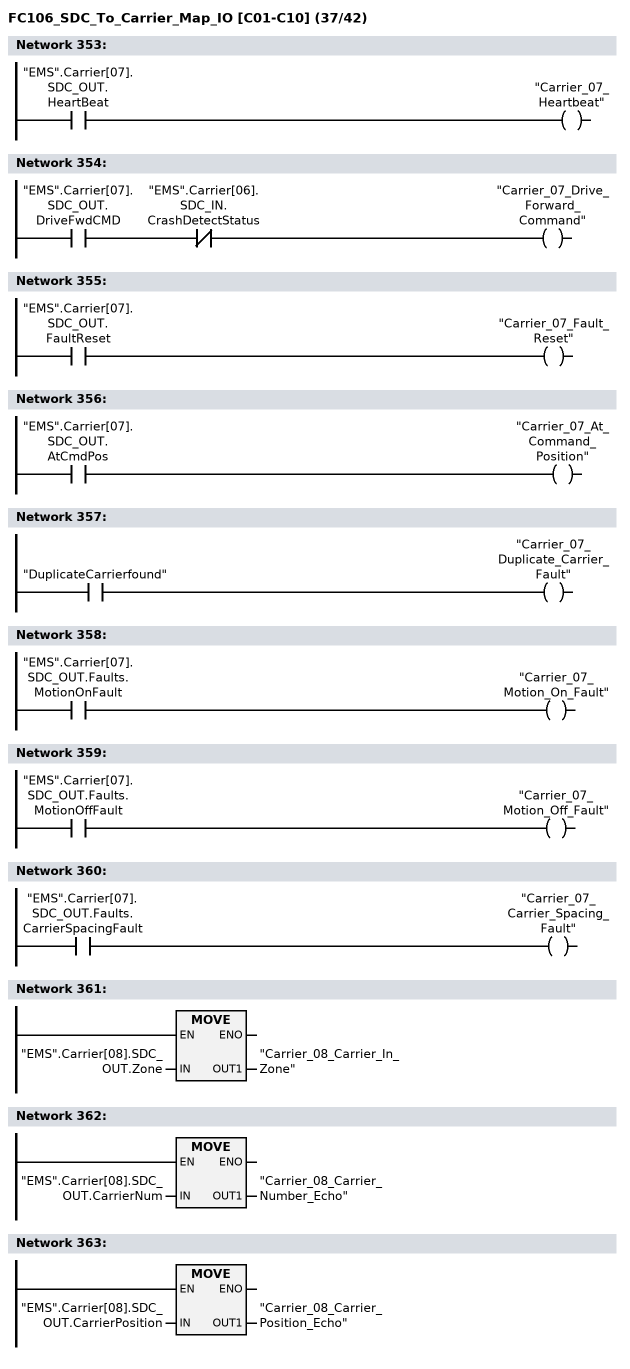
   RUNG wire#powerrail
      Contact( "EMS".Carrier[07].SDC_OUT.HeartBeat )
      Coil( "Carrier_07_Heartbeat" )
   END_RUNG
   // the same network as SCL:
   "Carrier_07_Heartbeat" := "EMS".Carrier[07].SDC_OUT.HeartBeat;
END_REGION

REGION Network 354
   RUNG wire#powerrail
      Contact( "EMS".Carrier[07].SDC_OUT.DriveFwdCMD )
      I_Contact( "EMS".Carrier[06].SDC_IN.CrashDetectStatus )
      Coil( "Carrier_07_Drive_Forward_Command" )
   END_RUNG
   // the same network as SCL:
   "Carrier_07_Drive_Forward_Command" := "EMS".Carrier[07].SDC_OUT.DriveFwdCMD AND NOT "EMS".Carrier[06].SDC_IN.CrashDetectStatus;
END_REGION

REGION Network 355
   RUNG wire#powerrail
      Contact( "EMS".Carrier[07].SDC_OUT.FaultReset )
      Coil( "Carrier_07_Fault_Reset" )
   END_RUNG
   // the same network as SCL:
   "Carrier_07_Fault_Reset" := "EMS".Carrier[07].SDC_OUT.FaultReset;
END_REGION

REGION Network 356
   RUNG wire#powerrail
      Contact( "EMS".Carrier[07].SDC_OUT.AtCmdPos )
      Coil( "Carrier_07_At_Command_Position" )
   END_RUNG
   // the same network as SCL:
   "Carrier_07_At_Command_Position" := "EMS".Carrier[07].SDC_OUT.AtCmdPos;
END_REGION

REGION Network 357
   RUNG wire#powerrail
      Contact( "DuplicateCarrierfound" )
      Coil( "Carrier_07_Duplicate_Carrier_Fault" )
   END_RUNG
   // the same network as SCL:
   "Carrier_07_Duplicate_Carrier_Fault" := "DuplicateCarrierfound";
END_REGION

REGION Network 358
   RUNG wire#powerrail
      Contact( "EMS".Carrier[07].SDC_OUT.Faults.MotionOnFault )
      Coil( "Carrier_07_Motion_On_Fault" )
   END_RUNG
   // the same network as SCL:
   "Carrier_07_Motion_On_Fault" := "EMS".Carrier[07].SDC_OUT.Faults.MotionOnFault;
END_REGION

REGION Network 359
   RUNG wire#powerrail
      Contact( "EMS".Carrier[07].SDC_OUT.Faults.MotionOffFault )
      Coil( "Carrier_07_Motion_Off_Fault" )
   END_RUNG
   // the same network as SCL:
   "Carrier_07_Motion_Off_Fault" := "EMS".Carrier[07].SDC_OUT.Faults.MotionOffFault;
END_REGION

REGION Network 360
   RUNG wire#powerrail
      Contact( "EMS".Carrier[07].SDC_OUT.Faults.CarrierSpacingFault )
      Coil( "Carrier_07_Carrier_Spacing_Fault" )
   END_RUNG
   // the same network as SCL:
   "Carrier_07_Carrier_Spacing_Fault" := "EMS".Carrier[07].SDC_OUT.Faults.CarrierSpacingFault;
END_REGION

REGION Network 361
   RUNG wire#powerrail
      Move(in := "EMS".Carrier[08].SDC_OUT.Zone, out1 => "Carrier_08_Carrier_In_Zone")
   END_RUNG
   // the same network as SCL:
   "Carrier_08_Carrier_In_Zone" := "EMS".Carrier[08].SDC_OUT.Zone;
END_REGION

REGION Network 362
   RUNG wire#powerrail
      Move(in := "EMS".Carrier[08].SDC_OUT.CarrierNum, out1 => "Carrier_08_Carrier_Number_Echo")
   END_RUNG
   // the same network as SCL:
   "Carrier_08_Carrier_Number_Echo" := "EMS".Carrier[08].SDC_OUT.CarrierNum;
END_REGION

REGION Network 363
   RUNG wire#powerrail
      Move(in := "EMS".Carrier[08].SDC_OUT.CarrierPosition, out1 => "Carrier_08_Carrier_Position_Echo")
   END_RUNG
   // the same network as SCL:
   "Carrier_08_Carrier_Position_Echo" := "EMS".Carrier[08].SDC_OUT.CarrierPosition;
END_REGION

REGION Network 364
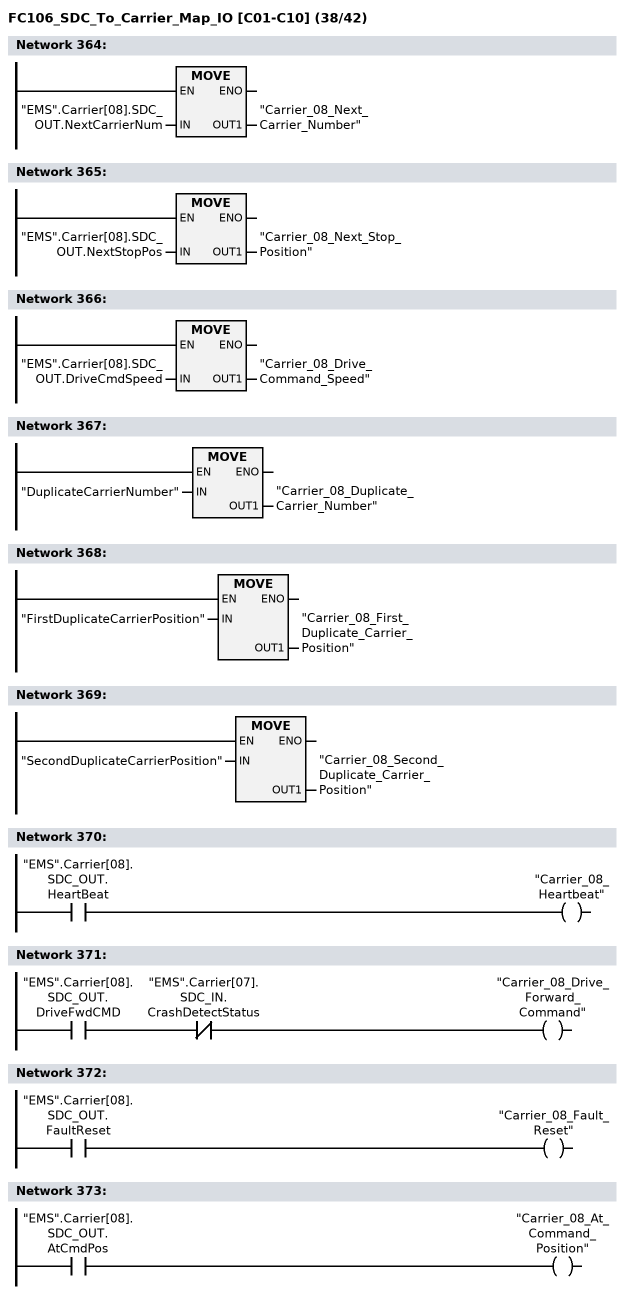
   RUNG wire#powerrail
      Move(in := "EMS".Carrier[08].SDC_OUT.NextCarrierNum, out1 => "Carrier_08_Next_Carrier_Number")
   END_RUNG
   // the same network as SCL:
   "Carrier_08_Next_Carrier_Number" := "EMS".Carrier[08].SDC_OUT.NextCarrierNum;
END_REGION

REGION Network 365
   RUNG wire#powerrail
      Move(in := "EMS".Carrier[08].SDC_OUT.NextStopPos, out1 => "Carrier_08_Next_Stop_Position")
   END_RUNG
   // the same network as SCL:
   "Carrier_08_Next_Stop_Position" := "EMS".Carrier[08].SDC_OUT.NextStopPos;
END_REGION

REGION Network 366
   RUNG wire#powerrail
      Move(in := "EMS".Carrier[08].SDC_OUT.DriveCmdSpeed, out1 => "Carrier_08_Drive_Command_Speed")
   END_RUNG
   // the same network as SCL:
   "Carrier_08_Drive_Command_Speed" := "EMS".Carrier[08].SDC_OUT.DriveCmdSpeed;
END_REGION

REGION Network 367
   RUNG wire#powerrail
      Move(in := "DuplicateCarrierNumber", out1 => "Carrier_08_Duplicate_Carrier_Number")
   END_RUNG
   // the same network as SCL:
   "Carrier_08_Duplicate_Carrier_Number" := "DuplicateCarrierNumber";
END_REGION

REGION Network 368
   RUNG wire#powerrail
      Move(in := "FirstDuplicateCarrierPosition", out1 => "Carrier_08_First_Duplicate_Carrier_Position")
   END_RUNG
   // the same network as SCL:
   "Carrier_08_First_Duplicate_Carrier_Position" := "FirstDuplicateCarrierPosition";
END_REGION

REGION Network 369
   RUNG wire#powerrail
      Move(in := "SecondDuplicateCarrierPosition", out1 => "Carrier_08_Second_Duplicate_Carrier_Position")
   END_RUNG
   // the same network as SCL:
   "Carrier_08_Second_Duplicate_Carrier_Position" := "SecondDuplicateCarrierPosition";
END_REGION

REGION Network 370
   RUNG wire#powerrail
      Contact( "EMS".Carrier[08].SDC_OUT.HeartBeat )
      Coil( "Carrier_08_Heartbeat" )
   END_RUNG
   // the same network as SCL:
   "Carrier_08_Heartbeat" := "EMS".Carrier[08].SDC_OUT.HeartBeat;
END_REGION

REGION Network 371
   RUNG wire#powerrail
      Contact( "EMS".Carrier[08].SDC_OUT.DriveFwdCMD )
      I_Contact( "EMS".Carrier[07].SDC_IN.CrashDetectStatus )
      Coil( "Carrier_08_Drive_Forward_Command" )
   END_RUNG
   // the same network as SCL:
   "Carrier_08_Drive_Forward_Command" := "EMS".Carrier[08].SDC_OUT.DriveFwdCMD AND NOT "EMS".Carrier[07].SDC_IN.CrashDetectStatus;
END_REGION

REGION Network 372
   RUNG wire#powerrail
      Contact( "EMS".Carrier[08].SDC_OUT.FaultReset )
      Coil( "Carrier_08_Fault_Reset" )
   END_RUNG
   // the same network as SCL:
   "Carrier_08_Fault_Reset" := "EMS".Carrier[08].SDC_OUT.FaultReset;
END_REGION

REGION Network 373
   RUNG wire#powerrail
      Contact( "EMS".Carrier[08].SDC_OUT.AtCmdPos )
      Coil( "Carrier_08_At_Command_Position" )
   END_RUNG
   // the same network as SCL:
   "Carrier_08_At_Command_Position" := "EMS".Carrier[08].SDC_OUT.AtCmdPos;
END_REGION

REGION Network 374
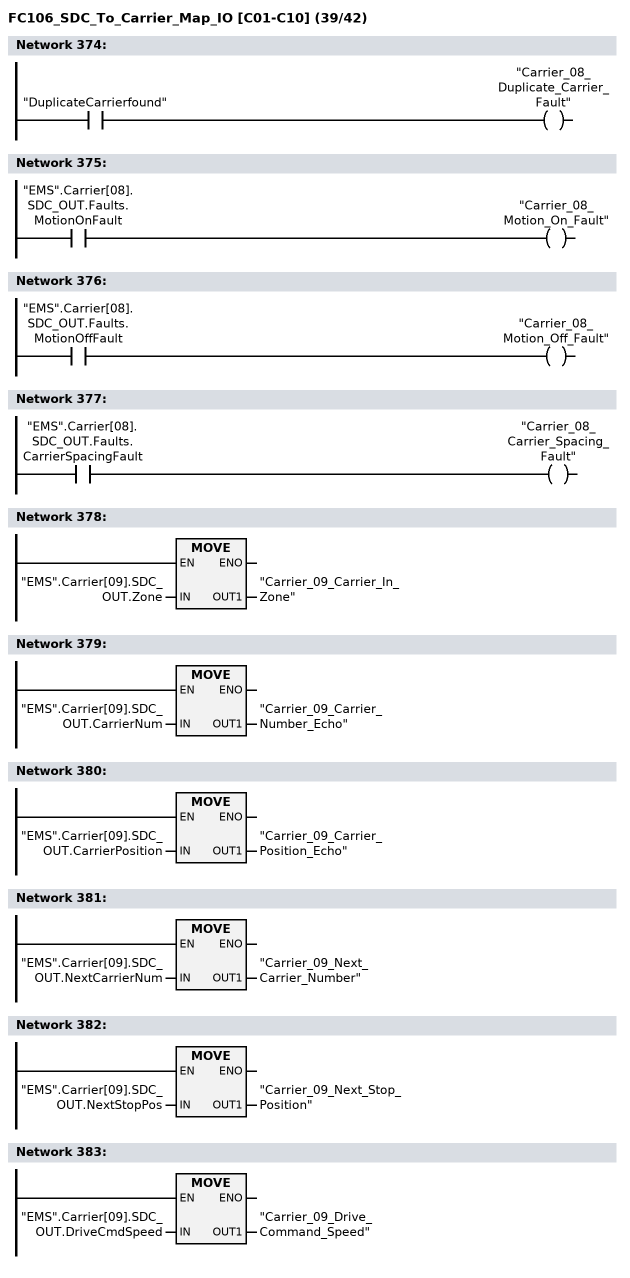
   RUNG wire#powerrail
      Contact( "DuplicateCarrierfound" )
      Coil( "Carrier_08_Duplicate_Carrier_Fault" )
   END_RUNG
   // the same network as SCL:
   "Carrier_08_Duplicate_Carrier_Fault" := "DuplicateCarrierfound";
END_REGION

REGION Network 375
   RUNG wire#powerrail
      Contact( "EMS".Carrier[08].SDC_OUT.Faults.MotionOnFault )
      Coil( "Carrier_08_Motion_On_Fault" )
   END_RUNG
   // the same network as SCL:
   "Carrier_08_Motion_On_Fault" := "EMS".Carrier[08].SDC_OUT.Faults.MotionOnFault;
END_REGION

REGION Network 376
   RUNG wire#powerrail
      Contact( "EMS".Carrier[08].SDC_OUT.Faults.MotionOffFault )
      Coil( "Carrier_08_Motion_Off_Fault" )
   END_RUNG
   // the same network as SCL:
   "Carrier_08_Motion_Off_Fault" := "EMS".Carrier[08].SDC_OUT.Faults.MotionOffFault;
END_REGION

REGION Network 377
   RUNG wire#powerrail
      Contact( "EMS".Carrier[08].SDC_OUT.Faults.CarrierSpacingFault )
      Coil( "Carrier_08_Carrier_Spacing_Fault" )
   END_RUNG
   // the same network as SCL:
   "Carrier_08_Carrier_Spacing_Fault" := "EMS".Carrier[08].SDC_OUT.Faults.CarrierSpacingFault;
END_REGION

REGION Network 378
   RUNG wire#powerrail
      Move(in := "EMS".Carrier[09].SDC_OUT.Zone, out1 => "Carrier_09_Carrier_In_Zone")
   END_RUNG
   // the same network as SCL:
   "Carrier_09_Carrier_In_Zone" := "EMS".Carrier[09].SDC_OUT.Zone;
END_REGION

REGION Network 379
   RUNG wire#powerrail
      Move(in := "EMS".Carrier[09].SDC_OUT.CarrierNum, out1 => "Carrier_09_Carrier_Number_Echo")
   END_RUNG
   // the same network as SCL:
   "Carrier_09_Carrier_Number_Echo" := "EMS".Carrier[09].SDC_OUT.CarrierNum;
END_REGION

REGION Network 380
   RUNG wire#powerrail
      Move(in := "EMS".Carrier[09].SDC_OUT.CarrierPosition, out1 => "Carrier_09_Carrier_Position_Echo")
   END_RUNG
   // the same network as SCL:
   "Carrier_09_Carrier_Position_Echo" := "EMS".Carrier[09].SDC_OUT.CarrierPosition;
END_REGION

REGION Network 381
   RUNG wire#powerrail
      Move(in := "EMS".Carrier[09].SDC_OUT.NextCarrierNum, out1 => "Carrier_09_Next_Carrier_Number")
   END_RUNG
   // the same network as SCL:
   "Carrier_09_Next_Carrier_Number" := "EMS".Carrier[09].SDC_OUT.NextCarrierNum;
END_REGION

REGION Network 382
   RUNG wire#powerrail
      Move(in := "EMS".Carrier[09].SDC_OUT.NextStopPos, out1 => "Carrier_09_Next_Stop_Position")
   END_RUNG
   // the same network as SCL:
   "Carrier_09_Next_Stop_Position" := "EMS".Carrier[09].SDC_OUT.NextStopPos;
END_REGION

REGION Network 383
   RUNG wire#powerrail
      Move(in := "EMS".Carrier[09].SDC_OUT.DriveCmdSpeed, out1 => "Carrier_09_Drive_Command_Speed")
   END_RUNG
   // the same network as SCL:
   "Carrier_09_Drive_Command_Speed" := "EMS".Carrier[09].SDC_OUT.DriveCmdSpeed;
END_REGION

REGION Network 384
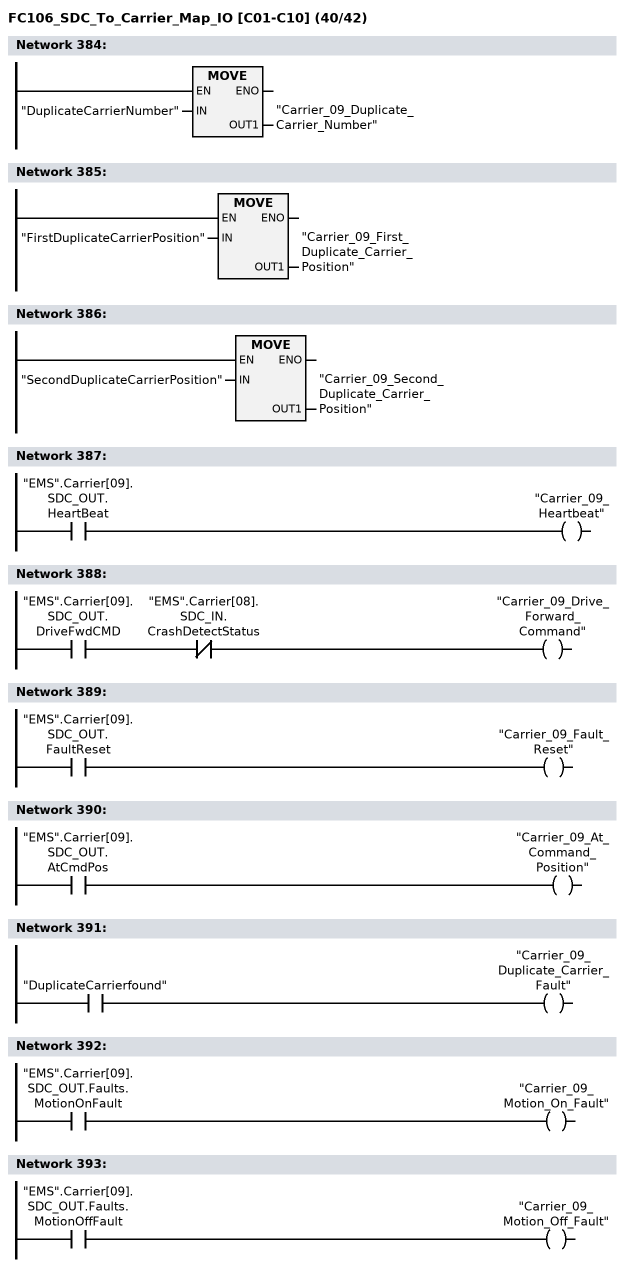
   RUNG wire#powerrail
      Move(in := "DuplicateCarrierNumber", out1 => "Carrier_09_Duplicate_Carrier_Number")
   END_RUNG
   // the same network as SCL:
   "Carrier_09_Duplicate_Carrier_Number" := "DuplicateCarrierNumber";
END_REGION

REGION Network 385
   RUNG wire#powerrail
      Move(in := "FirstDuplicateCarrierPosition", out1 => "Carrier_09_First_Duplicate_Carrier_Position")
   END_RUNG
   // the same network as SCL:
   "Carrier_09_First_Duplicate_Carrier_Position" := "FirstDuplicateCarrierPosition";
END_REGION

REGION Network 386
   RUNG wire#powerrail
      Move(in := "SecondDuplicateCarrierPosition", out1 => "Carrier_09_Second_Duplicate_Carrier_Position")
   END_RUNG
   // the same network as SCL:
   "Carrier_09_Second_Duplicate_Carrier_Position" := "SecondDuplicateCarrierPosition";
END_REGION

REGION Network 387
   RUNG wire#powerrail
      Contact( "EMS".Carrier[09].SDC_OUT.HeartBeat )
      Coil( "Carrier_09_Heartbeat" )
   END_RUNG
   // the same network as SCL:
   "Carrier_09_Heartbeat" := "EMS".Carrier[09].SDC_OUT.HeartBeat;
END_REGION

REGION Network 388
   RUNG wire#powerrail
      Contact( "EMS".Carrier[09].SDC_OUT.DriveFwdCMD )
      I_Contact( "EMS".Carrier[08].SDC_IN.CrashDetectStatus )
      Coil( "Carrier_09_Drive_Forward_Command" )
   END_RUNG
   // the same network as SCL:
   "Carrier_09_Drive_Forward_Command" := "EMS".Carrier[09].SDC_OUT.DriveFwdCMD AND NOT "EMS".Carrier[08].SDC_IN.CrashDetectStatus;
END_REGION

REGION Network 389
   RUNG wire#powerrail
      Contact( "EMS".Carrier[09].SDC_OUT.FaultReset )
      Coil( "Carrier_09_Fault_Reset" )
   END_RUNG
   // the same network as SCL:
   "Carrier_09_Fault_Reset" := "EMS".Carrier[09].SDC_OUT.FaultReset;
END_REGION

REGION Network 390
   RUNG wire#powerrail
      Contact( "EMS".Carrier[09].SDC_OUT.AtCmdPos )
      Coil( "Carrier_09_At_Command_Position" )
   END_RUNG
   // the same network as SCL:
   "Carrier_09_At_Command_Position" := "EMS".Carrier[09].SDC_OUT.AtCmdPos;
END_REGION

REGION Network 391
   RUNG wire#powerrail
      Contact( "DuplicateCarrierfound" )
      Coil( "Carrier_09_Duplicate_Carrier_Fault" )
   END_RUNG
   // the same network as SCL:
   "Carrier_09_Duplicate_Carrier_Fault" := "DuplicateCarrierfound";
END_REGION

REGION Network 392
   RUNG wire#powerrail
      Contact( "EMS".Carrier[09].SDC_OUT.Faults.MotionOnFault )
      Coil( "Carrier_09_Motion_On_Fault" )
   END_RUNG
   // the same network as SCL:
   "Carrier_09_Motion_On_Fault" := "EMS".Carrier[09].SDC_OUT.Faults.MotionOnFault;
END_REGION

REGION Network 393
   RUNG wire#powerrail
      Contact( "EMS".Carrier[09].SDC_OUT.Faults.MotionOffFault )
      Coil( "Carrier_09_Motion_Off_Fault" )
   END_RUNG
   // the same network as SCL:
   "Carrier_09_Motion_Off_Fault" := "EMS".Carrier[09].SDC_OUT.Faults.MotionOffFault;
END_REGION

REGION Network 394
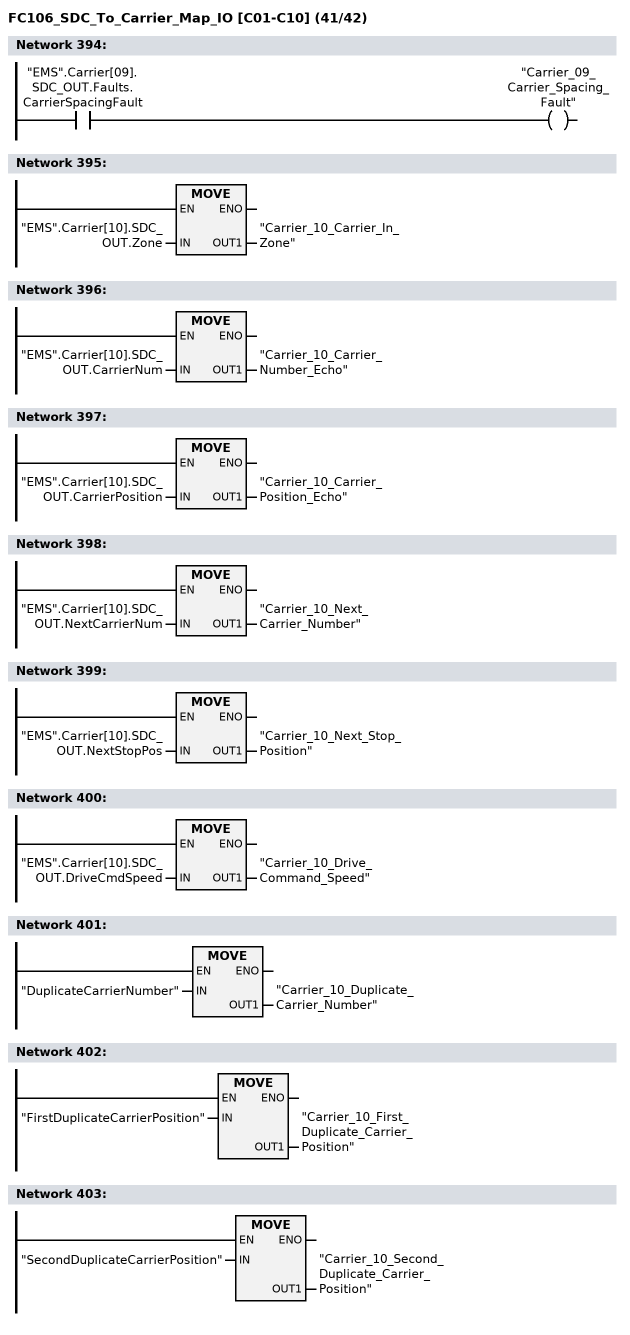
   RUNG wire#powerrail
      Contact( "EMS".Carrier[09].SDC_OUT.Faults.CarrierSpacingFault )
      Coil( "Carrier_09_Carrier_Spacing_Fault" )
   END_RUNG
   // the same network as SCL:
   "Carrier_09_Carrier_Spacing_Fault" := "EMS".Carrier[09].SDC_OUT.Faults.CarrierSpacingFault;
END_REGION

REGION Network 395
   RUNG wire#powerrail
      Move(in := "EMS".Carrier[10].SDC_OUT.Zone, out1 => "Carrier_10_Carrier_In_Zone")
   END_RUNG
   // the same network as SCL:
   "Carrier_10_Carrier_In_Zone" := "EMS".Carrier[10].SDC_OUT.Zone;
END_REGION

REGION Network 396
   RUNG wire#powerrail
      Move(in := "EMS".Carrier[10].SDC_OUT.CarrierNum, out1 => "Carrier_10_Carrier_Number_Echo")
   END_RUNG
   // the same network as SCL:
   "Carrier_10_Carrier_Number_Echo" := "EMS".Carrier[10].SDC_OUT.CarrierNum;
END_REGION

REGION Network 397
   RUNG wire#powerrail
      Move(in := "EMS".Carrier[10].SDC_OUT.CarrierPosition, out1 => "Carrier_10_Carrier_Position_Echo")
   END_RUNG
   // the same network as SCL:
   "Carrier_10_Carrier_Position_Echo" := "EMS".Carrier[10].SDC_OUT.CarrierPosition;
END_REGION

REGION Network 398
   RUNG wire#powerrail
      Move(in := "EMS".Carrier[10].SDC_OUT.NextCarrierNum, out1 => "Carrier_10_Next_Carrier_Number")
   END_RUNG
   // the same network as SCL:
   "Carrier_10_Next_Carrier_Number" := "EMS".Carrier[10].SDC_OUT.NextCarrierNum;
END_REGION

REGION Network 399
   RUNG wire#powerrail
      Move(in := "EMS".Carrier[10].SDC_OUT.NextStopPos, out1 => "Carrier_10_Next_Stop_Position")
   END_RUNG
   // the same network as SCL:
   "Carrier_10_Next_Stop_Position" := "EMS".Carrier[10].SDC_OUT.NextStopPos;
END_REGION

REGION Network 400
   RUNG wire#powerrail
      Move(in := "EMS".Carrier[10].SDC_OUT.DriveCmdSpeed, out1 => "Carrier_10_Drive_Command_Speed")
   END_RUNG
   // the same network as SCL:
   "Carrier_10_Drive_Command_Speed" := "EMS".Carrier[10].SDC_OUT.DriveCmdSpeed;
END_REGION

REGION Network 401
   RUNG wire#powerrail
      Move(in := "DuplicateCarrierNumber", out1 => "Carrier_10_Duplicate_Carrier_Number")
   END_RUNG
   // the same network as SCL:
   "Carrier_10_Duplicate_Carrier_Number" := "DuplicateCarrierNumber";
END_REGION

REGION Network 402
   RUNG wire#powerrail
      Move(in := "FirstDuplicateCarrierPosition", out1 => "Carrier_10_First_Duplicate_Carrier_Position")
   END_RUNG
   // the same network as SCL:
   "Carrier_10_First_Duplicate_Carrier_Position" := "FirstDuplicateCarrierPosition";
END_REGION

REGION Network 403
   RUNG wire#powerrail
      Move(in := "SecondDuplicateCarrierPosition", out1 => "Carrier_10_Second_Duplicate_Carrier_Position")
   END_RUNG
   // the same network as SCL:
   "Carrier_10_Second_Duplicate_Carrier_Position" := "SecondDuplicateCarrierPosition";
END_REGION

REGION Network 404
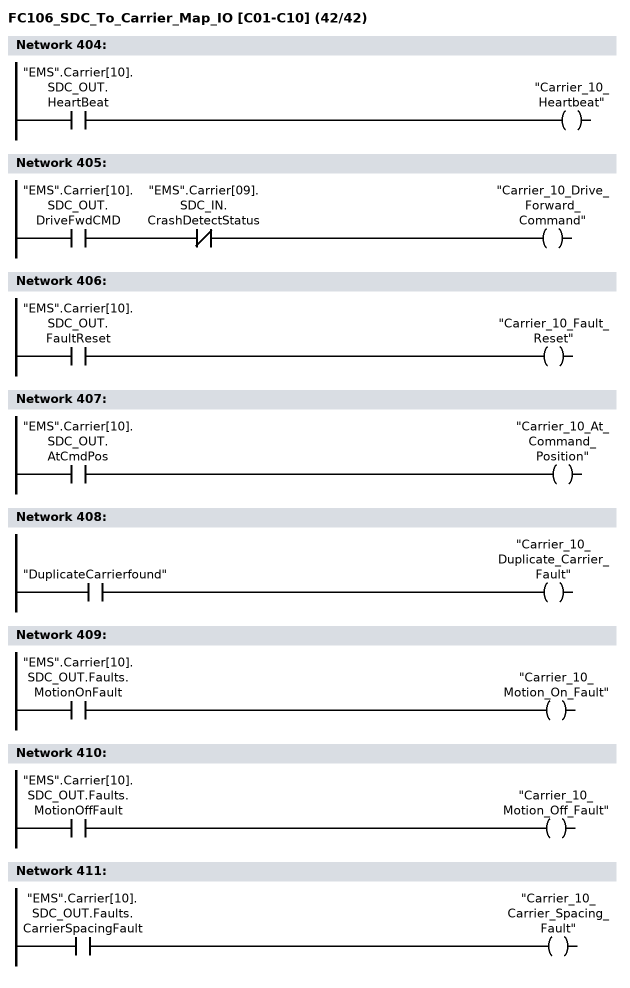
   RUNG wire#powerrail
      Contact( "EMS".Carrier[10].SDC_OUT.HeartBeat )
      Coil( "Carrier_10_Heartbeat" )
   END_RUNG
   // the same network as SCL:
   "Carrier_10_Heartbeat" := "EMS".Carrier[10].SDC_OUT.HeartBeat;
END_REGION

REGION Network 405
   RUNG wire#powerrail
      Contact( "EMS".Carrier[10].SDC_OUT.DriveFwdCMD )
      I_Contact( "EMS".Carrier[09].SDC_IN.CrashDetectStatus )
      Coil( "Carrier_10_Drive_Forward_Command" )
   END_RUNG
   // the same network as SCL:
   "Carrier_10_Drive_Forward_Command" := "EMS".Carrier[10].SDC_OUT.DriveFwdCMD AND NOT "EMS".Carrier[09].SDC_IN.CrashDetectStatus;
END_REGION

REGION Network 406
   RUNG wire#powerrail
      Contact( "EMS".Carrier[10].SDC_OUT.FaultReset )
      Coil( "Carrier_10_Fault_Reset" )
   END_RUNG
   // the same network as SCL:
   "Carrier_10_Fault_Reset" := "EMS".Carrier[10].SDC_OUT.FaultReset;
END_REGION

REGION Network 407
   RUNG wire#powerrail
      Contact( "EMS".Carrier[10].SDC_OUT.AtCmdPos )
      Coil( "Carrier_10_At_Command_Position" )
   END_RUNG
   // the same network as SCL:
   "Carrier_10_At_Command_Position" := "EMS".Carrier[10].SDC_OUT.AtCmdPos;
END_REGION

REGION Network 408
   RUNG wire#powerrail
      Contact( "DuplicateCarrierfound" )
      Coil( "Carrier_10_Duplicate_Carrier_Fault" )
   END_RUNG
   // the same network as SCL:
   "Carrier_10_Duplicate_Carrier_Fault" := "DuplicateCarrierfound";
END_REGION

REGION Network 409
   RUNG wire#powerrail
      Contact( "EMS".Carrier[10].SDC_OUT.Faults.MotionOnFault )
      Coil( "Carrier_10_Motion_On_Fault" )
   END_RUNG
   // the same network as SCL:
   "Carrier_10_Motion_On_Fault" := "EMS".Carrier[10].SDC_OUT.Faults.MotionOnFault;
END_REGION

REGION Network 410
   RUNG wire#powerrail
      Contact( "EMS".Carrier[10].SDC_OUT.Faults.MotionOffFault )
      Coil( "Carrier_10_Motion_Off_Fault" )
   END_RUNG
   // the same network as SCL:
   "Carrier_10_Motion_Off_Fault" := "EMS".Carrier[10].SDC_OUT.Faults.MotionOffFault;
END_REGION

REGION Network 411
   RUNG wire#powerrail
      Contact( "EMS".Carrier[10].SDC_OUT.Faults.CarrierSpacingFault )
      Coil( "Carrier_10_Carrier_Spacing_Fault" )
   END_RUNG
   // the same network as SCL:
   "Carrier_10_Carrier_Spacing_Fault" := "EMS".Carrier[10].SDC_OUT.Faults.CarrierSpacingFault;
END_REGION
END_FUNCTION

FUNCTION "FC107_SDC_To_Carrier_Map_IO [C11-C20]" : Void   // FC107, LAD
{ S7_Optimized_Access := 'TRUE' }
VERSION : 0.1
BEGIN

REGION Network 1
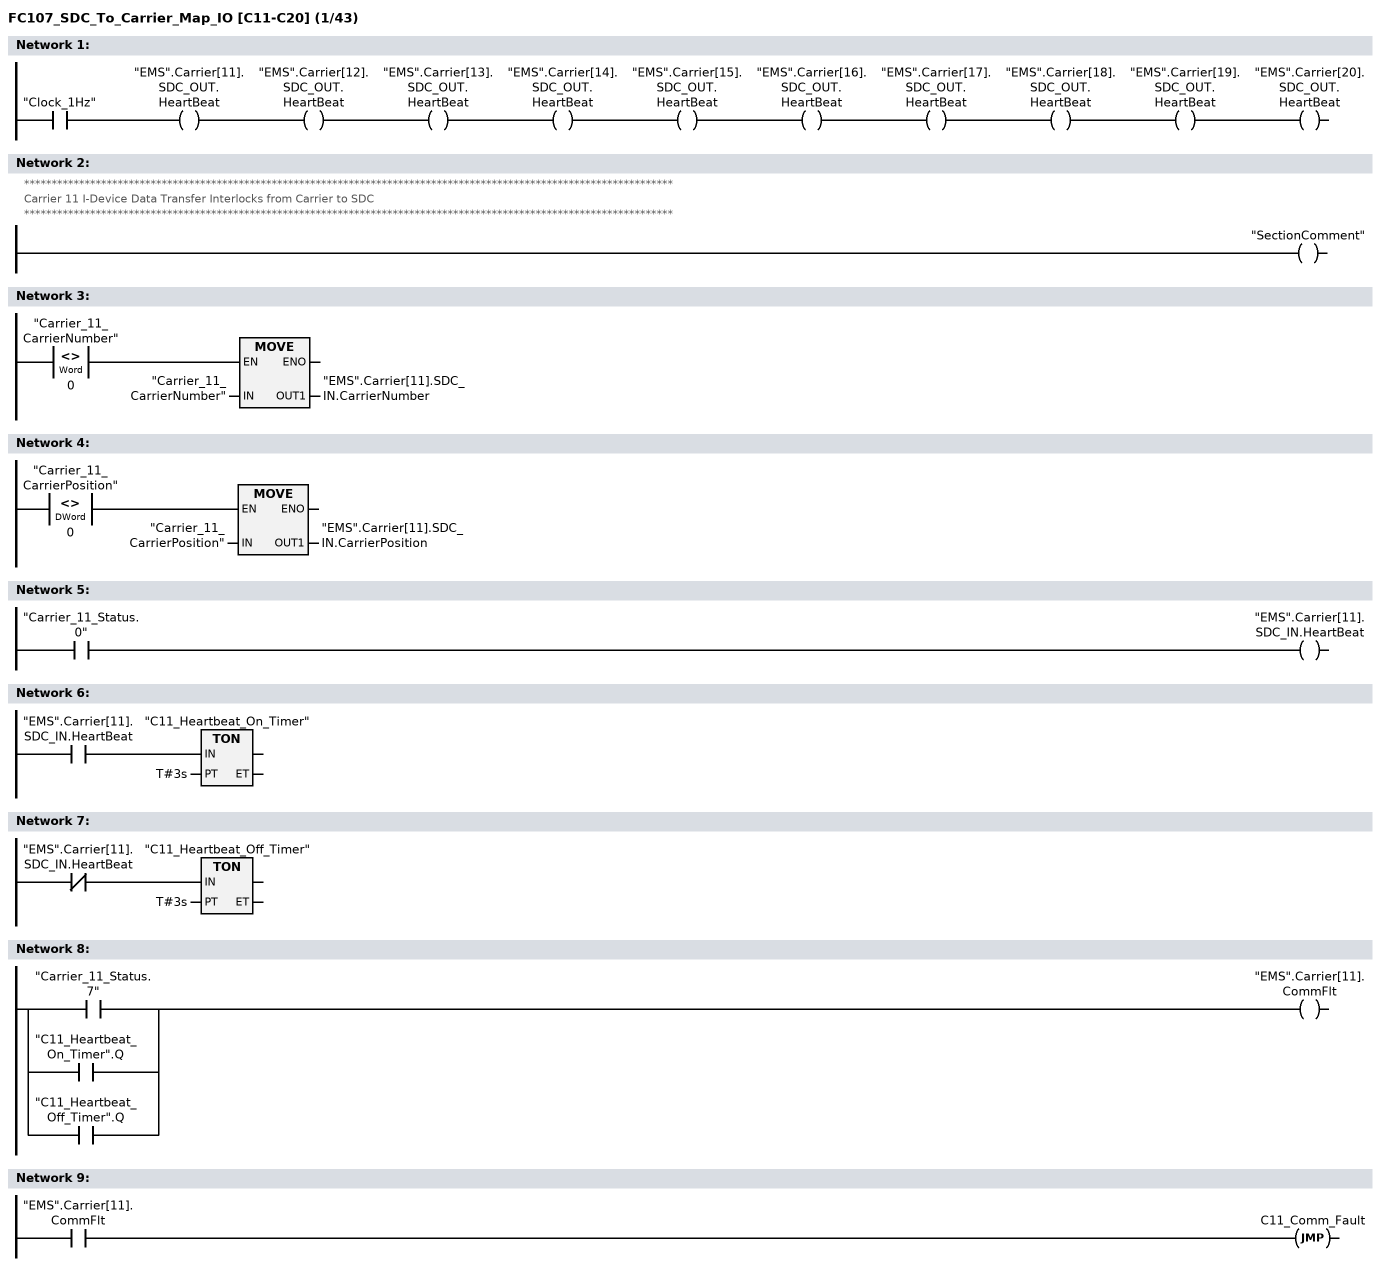
   RUNG wire#powerrail
      Contact( "Clock_1Hz" )
      Coil( "EMS".Carrier[11].SDC_OUT.HeartBeat )
      Coil( "EMS".Carrier[12].SDC_OUT.HeartBeat )
      Coil( "EMS".Carrier[13].SDC_OUT.HeartBeat )
      Coil( "EMS".Carrier[14].SDC_OUT.HeartBeat )
      Coil( "EMS".Carrier[15].SDC_OUT.HeartBeat )
      Coil( "EMS".Carrier[16].SDC_OUT.HeartBeat )
      Coil( "EMS".Carrier[17].SDC_OUT.HeartBeat )
      Coil( "EMS".Carrier[18].SDC_OUT.HeartBeat )
      Coil( "EMS".Carrier[19].SDC_OUT.HeartBeat )
      Coil( "EMS".Carrier[20].SDC_OUT.HeartBeat )
   END_RUNG
   // the same network as SCL:
   "EMS".Carrier[11].SDC_OUT.HeartBeat := "Clock_1Hz";
   "EMS".Carrier[12].SDC_OUT.HeartBeat := "Clock_1Hz";
   "EMS".Carrier[13].SDC_OUT.HeartBeat := "Clock_1Hz";
   "EMS".Carrier[14].SDC_OUT.HeartBeat := "Clock_1Hz";
   "EMS".Carrier[15].SDC_OUT.HeartBeat := "Clock_1Hz";
   "EMS".Carrier[16].SDC_OUT.HeartBeat := "Clock_1Hz";
   "EMS".Carrier[17].SDC_OUT.HeartBeat := "Clock_1Hz";
   "EMS".Carrier[18].SDC_OUT.HeartBeat := "Clock_1Hz";
   "EMS".Carrier[19].SDC_OUT.HeartBeat := "Clock_1Hz";
   "EMS".Carrier[20].SDC_OUT.HeartBeat := "Clock_1Hz";
END_REGION

REGION Network 2
   // **********************************************************************************************************************
   // 
   // Carrier 11 I-Device Data Transfer Interlocks from Carrier to SDC
   // 
   // **********************************************************************************************************************
   RUNG wire#powerrail
      Coil( "SectionComment" )
   END_RUNG
   // the same network as SCL:
   "SectionComment" := TRUE;
END_REGION

REGION Network 3
   RUNG wire#powerrail
      { S7_Templates := "SrcType := Word" } NE_Contact(in1 := "Carrier_11_CarrierNumber", in2 := 0)
      Move(in := "Carrier_11_CarrierNumber", out1 => "EMS".Carrier[11].SDC_IN.CarrierNumber)
   END_RUNG
   // the same network as SCL:
   IF "Carrier_11_CarrierNumber" <> 0 THEN
       "EMS".Carrier[11].SDC_IN.CarrierNumber := "Carrier_11_CarrierNumber";
   END_IF;
END_REGION

REGION Network 4
   RUNG wire#powerrail
      { S7_Templates := "SrcType := DWord" } NE_Contact(in1 := "Carrier_11_CarrierPosition", in2 := 0)
      Move(in := "Carrier_11_CarrierPosition", out1 => "EMS".Carrier[11].SDC_IN.CarrierPosition)
   END_RUNG
   // the same network as SCL:
   IF "Carrier_11_CarrierPosition" <> 0 THEN
       "EMS".Carrier[11].SDC_IN.CarrierPosition := "Carrier_11_CarrierPosition";
   END_IF;
END_REGION

REGION Network 5
   RUNG wire#powerrail
      Contact( "Carrier_11_Status.0" )
      Coil( "EMS".Carrier[11].SDC_IN.HeartBeat )
   END_RUNG
   // the same network as SCL:
   "EMS".Carrier[11].SDC_IN.HeartBeat := "Carrier_11_Status.0";
END_REGION

REGION Network 6
   "C11_Heartbeat_On_Timer".TON(IN := "EMS".Carrier[11].SDC_IN.HeartBeat, PT := T#3s);
END_REGION

REGION Network 7
   "C11_Heartbeat_Off_Timer".TON(IN := NOT "EMS".Carrier[11].SDC_IN.HeartBeat, PT := T#3s);
END_REGION

REGION Network 8
   RUNG wire#powerrail
      Contact( "Carrier_11_Status.7" )
      wire#w1
      Coil( "EMS".Carrier[11].CommFlt )
   END_RUNG
   RUNG wire#powerrail
      Contact( "C11_Heartbeat_On_Timer".Q )
   END_RUNG wire#w1
   RUNG wire#powerrail
      Contact( "C11_Heartbeat_Off_Timer".Q )
   END_RUNG wire#w1
   // the same network as SCL:
   "EMS".Carrier[11].CommFlt := "Carrier_11_Status.7" OR "C11_Heartbeat_On_Timer".Q OR "C11_Heartbeat_Off_Timer".Q;
END_REGION

REGION Network 9
   RUNG wire#powerrail
      Contact( "EMS".Carrier[11].CommFlt )
      JumpCoil( C11_Comm_Fault )
   END_RUNG
   // the same network as SCL:
   IF "EMS".Carrier[11].CommFlt THEN GOTO C11_Comm_Fault; END_IF;
END_REGION

REGION Network 10
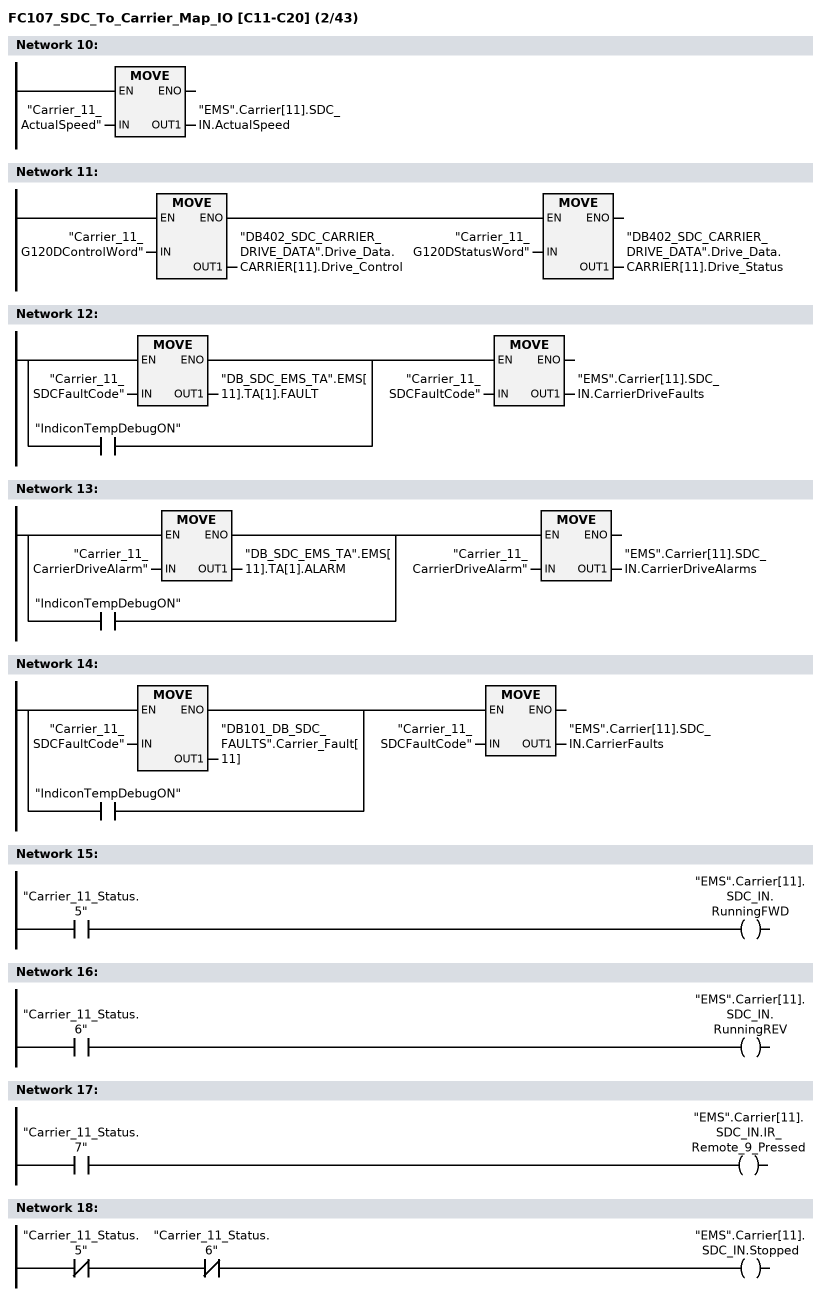
   RUNG wire#powerrail
      Move(in := "Carrier_11_ActualSpeed", out1 => "EMS".Carrier[11].SDC_IN.ActualSpeed)
   END_RUNG
   // the same network as SCL:
   "EMS".Carrier[11].SDC_IN.ActualSpeed := "Carrier_11_ActualSpeed";
END_REGION

REGION Network 11
   RUNG wire#powerrail
      Move(in := "Carrier_11_G120DControlWord", out1 => "DB402_SDC_CARRIER_DRIVE_DATA".Drive_Data.CARRIER[11].Drive_Control)
      Move(in := "Carrier_11_G120DStatusWord", out1 => "DB402_SDC_CARRIER_DRIVE_DATA".Drive_Data.CARRIER[11].Drive_Status)
   END_RUNG
   // the same network as SCL:
   "DB402_SDC_CARRIER_DRIVE_DATA".Drive_Data.CARRIER[11].Drive_Control := "Carrier_11_G120DControlWord";
   "DB402_SDC_CARRIER_DRIVE_DATA".Drive_Data.CARRIER[11].Drive_Status := "Carrier_11_G120DStatusWord";
END_REGION

REGION Network 12
   RUNG wire#powerrail
      Move(in := "Carrier_11_SDCFaultCode", out1 => "DB_SDC_EMS_TA".EMS[11].TA[1].FAULT)
      wire#w1
      Move(in := "Carrier_11_SDCFaultCode", out1 => "EMS".Carrier[11].SDC_IN.CarrierDriveFaults)
   END_RUNG
   RUNG wire#powerrail
      Contact( "IndiconTempDebugON" )
   END_RUNG wire#w1
   // the same network as SCL:
   "DB_SDC_EMS_TA".EMS[11].TA[1].FAULT := "Carrier_11_SDCFaultCode";
   IF TRUE OR "IndiconTempDebugON" THEN
       "EMS".Carrier[11].SDC_IN.CarrierDriveFaults := "Carrier_11_SDCFaultCode";
   END_IF;
END_REGION

REGION Network 13
   RUNG wire#powerrail
      Move(in := "Carrier_11_CarrierDriveAlarm", out1 => "DB_SDC_EMS_TA".EMS[11].TA[1].ALARM)
      wire#w1
      Move(in := "Carrier_11_CarrierDriveAlarm", out1 => "EMS".Carrier[11].SDC_IN.CarrierDriveAlarms)
   END_RUNG
   RUNG wire#powerrail
      Contact( "IndiconTempDebugON" )
   END_RUNG wire#w1
   // the same network as SCL:
   "DB_SDC_EMS_TA".EMS[11].TA[1].ALARM := "Carrier_11_CarrierDriveAlarm";
   IF TRUE OR "IndiconTempDebugON" THEN
       "EMS".Carrier[11].SDC_IN.CarrierDriveAlarms := "Carrier_11_CarrierDriveAlarm";
   END_IF;
END_REGION

REGION Network 14
   RUNG wire#powerrail
      Move(in := "Carrier_11_SDCFaultCode", out1 => "DB101_DB_SDC_FAULTS".Carrier_Fault[11])
      wire#w1
      Move(in := "Carrier_11_SDCFaultCode", out1 => "EMS".Carrier[11].SDC_IN.CarrierFaults)
   END_RUNG
   RUNG wire#powerrail
      Contact( "IndiconTempDebugON" )
   END_RUNG wire#w1
   // the same network as SCL:
   "DB101_DB_SDC_FAULTS".Carrier_Fault[11] := "Carrier_11_SDCFaultCode";
   IF TRUE OR "IndiconTempDebugON" THEN
       "EMS".Carrier[11].SDC_IN.CarrierFaults := "Carrier_11_SDCFaultCode";
   END_IF;
END_REGION

REGION Network 15
   RUNG wire#powerrail
      Contact( "Carrier_11_Status.5" )
      Coil( "EMS".Carrier[11].SDC_IN.RunningFWD )
   END_RUNG
   // the same network as SCL:
   "EMS".Carrier[11].SDC_IN.RunningFWD := "Carrier_11_Status.5";
END_REGION

REGION Network 16
   RUNG wire#powerrail
      Contact( "Carrier_11_Status.6" )
      Coil( "EMS".Carrier[11].SDC_IN.RunningREV )
   END_RUNG
   // the same network as SCL:
   "EMS".Carrier[11].SDC_IN.RunningREV := "Carrier_11_Status.6";
END_REGION

REGION Network 17
   RUNG wire#powerrail
      Contact( "Carrier_11_Status.7" )
      Coil( "EMS".Carrier[11].SDC_IN.IR_Remote_9_Pressed )
   END_RUNG
   // the same network as SCL:
   "EMS".Carrier[11].SDC_IN.IR_Remote_9_Pressed := "Carrier_11_Status.7";
END_REGION

REGION Network 18
   RUNG wire#powerrail
      I_Contact( "Carrier_11_Status.5" )
      I_Contact( "Carrier_11_Status.6" )
      Coil( "EMS".Carrier[11].SDC_IN.Stopped )
   END_RUNG
   // the same network as SCL:
   "EMS".Carrier[11].SDC_IN.Stopped := NOT "Carrier_11_Status.5" AND NOT "Carrier_11_Status.6";
END_REGION

REGION Network 19
